(* Logix 5000 project; controller OWF Emulate 5570 rev 30.12; software revision 30.00 *) (continued)
   	OWF_Key[105,2]:=1079186439;
   	OWF_Key[105,3]:=354175718;
   	OWF_Key[105,4]:=460014900;
   	OWF_Key[105,5]:=657327792;
   	OWF_Key[105,6]:=1238184223;
   	OWF_Key[105,7]:=613398807;
   	OWF_Key[105,8]:=313681701;
   	OWF_Key[106,0]:=623677644;
   	OWF_Key[106,1]:=1206586343;
   	OWF_Key[106,2]:=1211299162;
   	OWF_Key[106,3]:=1368157030;
   	OWF_Key[106,4]:=1726692177;
   	OWF_Key[106,5]:=909079139;
   	OWF_Key[106,6]:=1189133566;
   	OWF_Key[106,7]:=1775183384;
   	OWF_Key[106,8]:=1947314078;
   	OWF_Key[107,0]:=795842741;
   	OWF_Key[107,1]:=5243211;
   	OWF_Key[107,2]:=2117485737;
   	OWF_Key[107,3]:=1222955765;
   	OWF_Key[107,4]:=1010466652;
   	OWF_Key[107,5]:=1366757084;
   	OWF_Key[107,6]:=1745897474;
   	OWF_Key[107,7]:=1196628900;
   	OWF_Key[107,8]:=422811900;
   	OWF_Key[108,0]:=51546250;
   	OWF_Key[108,1]:=1371654065;
   	OWF_Key[108,2]:=594730613;
   	OWF_Key[108,3]:=1178928938;
   	OWF_Key[108,4]:=19658574;
   	OWF_Key[108,5]:=44268080;
   	OWF_Key[108,6]:=1705061822;
   	OWF_Key[108,7]:=765733996;
   	OWF_Key[108,8]:=254021521;
   	OWF_Key[109,0]:=1089931182;
   	OWF_Key[109,1]:=456261576;
   	OWF_Key[109,2]:=1032396223;
   	OWF_Key[109,3]:=1215239566;
   	OWF_Key[109,4]:=1432021362;
   	OWF_Key[109,5]:=1482695855;
   	OWF_Key[109,6]:=471826292;
   	OWF_Key[109,7]:=1639233209;
   	OWF_Key[109,8]:=33522508;
   	OWF_Key[110,0]:=1943548851;
   	OWF_Key[110,1]:=188222712;
   	OWF_Key[110,2]:=2073166455;
   	OWF_Key[110,3]:=1482931688;
   	OWF_Key[110,4]:=816300030;
   	OWF_Key[110,5]:=246963335;
   	OWF_Key[110,6]:=313723350;
   	OWF_Key[110,7]:=331932254;
   	OWF_Key[110,8]:=1039085928;
   	OWF_Key[111,0]:=913532003;
   	OWF_Key[111,1]:=1339665160;
   	OWF_Key[111,2]:=14150618;
   	OWF_Key[111,3]:=743204030;
   	OWF_Key[111,4]:=2083710274;
   	OWF_Key[111,5]:=1872451661;
   	OWF_Key[111,6]:=1349153003;
   	OWF_Key[111,7]:=373058060;
   	OWF_Key[111,8]:=778338392;
   	OWF_Key[112,0]:=1413062923;
   	OWF_Key[112,1]:=1525503190;
   	OWF_Key[112,2]:=153669953;
   	OWF_Key[112,3]:=1075488387;
   	OWF_Key[112,4]:=1611202824;
   	OWF_Key[112,5]:=842678039;
   	OWF_Key[112,6]:=1878241110;
   	OWF_Key[112,7]:=2094622845;
   	OWF_Key[112,8]:=346061363;
   	OWF_Key[113,0]:=2007662486;
   	OWF_Key[113,1]:=609926961;
   	OWF_Key[113,2]:=208768431;
   	OWF_Key[113,3]:=1089775410;
   	OWF_Key[113,4]:=2139360128;
   	OWF_Key[113,5]:=246842036;
   	OWF_Key[113,6]:=437887573;
   	OWF_Key[113,7]:=1715106097;
   	OWF_Key[113,8]:=1931243001;
   	OWF_Key[114,0]:=1695412974;
   	OWF_Key[114,1]:=75402688;
   	OWF_Key[114,2]:=1324107774;
   	OWF_Key[114,3]:=1762126149;
   	OWF_Key[114,4]:=2045453401;
   	OWF_Key[114,5]:=1322782179;
   	OWF_Key[114,6]:=560014314;
   	OWF_Key[114,7]:=113230679;
   	OWF_Key[114,8]:=1460013455;
   	OWF_Key[115,0]:=1522550142;
   	OWF_Key[115,1]:=181079064;
   	OWF_Key[115,2]:=1318356612;
   	OWF_Key[115,3]:=1089396761;
   	OWF_Key[115,4]:=2100774490;
   	OWF_Key[115,5]:=1187593175;
   	OWF_Key[115,6]:=673723015;
   	OWF_Key[115,7]:=1625716407;
   	OWF_Key[115,8]:=157879385;
   	OWF_Key[116,0]:=1574439302;
   	OWF_Key[116,1]:=1171649064;
   	OWF_Key[116,2]:=1725295889;
   	OWF_Key[116,3]:=1508609966;
   	OWF_Key[116,4]:=893053329;
   	OWF_Key[116,5]:=2022024439;
   	OWF_Key[116,6]:=1645938530;
   	OWF_Key[116,7]:=1690657533;
   	OWF_Key[116,8]:=1383145517;
   	OWF_Key[117,0]:=255569215;
   	OWF_Key[117,1]:=1987873809;
   	OWF_Key[117,2]:=397411303;
   	OWF_Key[117,3]:=1688889668;
   	OWF_Key[117,4]:=222285489;
   	OWF_Key[117,5]:=449962612;
   	OWF_Key[117,6]:=751498151;
   	OWF_Key[117,7]:=708509537;
   	OWF_Key[117,8]:=2068975187;
   	OWF_Key[118,0]:=755822791;
   	OWF_Key[118,1]:=705169811;
   	OWF_Key[118,2]:=1142286417;
   	OWF_Key[118,3]:=157784650;
   	OWF_Key[118,4]:=506439582;
   	OWF_Key[118,5]:=1051639190;
   	OWF_Key[118,6]:=1903419853;
   	OWF_Key[118,7]:=1851507373;
   	OWF_Key[118,8]:=1030591932;
   	OWF_Key[119,0]:=2057479898;
   	OWF_Key[119,1]:=2036906294;
   	OWF_Key[119,2]:=254059922;
   	OWF_Key[119,3]:=849168680;
   	OWF_Key[119,4]:=301288022;
   	OWF_Key[119,5]:=1586180160;
   	OWF_Key[119,6]:=434263535;
   	OWF_Key[119,7]:=1375534755;
   	OWF_Key[119,8]:=967855848;
   	OWF_Key[120,0]:=1790809297;
   	OWF_Key[120,1]:=913198018;
   	OWF_Key[120,2]:=996748500;
   	OWF_Key[120,3]:=326041118;
   	OWF_Key[120,4]:=1340890547;
   	OWF_Key[120,5]:=1923120038;
   	OWF_Key[120,6]:=122657393;
   	OWF_Key[120,7]:=1589302007;
   	OWF_Key[120,8]:=1782178774;
   	OWF_Key[121,0]:=82130336;
   	OWF_Key[121,1]:=1724730757;
   	OWF_Key[121,2]:=1991211720;
   	OWF_Key[121,3]:=559635139;
   	OWF_Key[121,4]:=1292994698;
   	OWF_Key[121,5]:=884899297;
   	OWF_Key[121,6]:=54837547;
   	OWF_Key[121,7]:=1512359967;
   	OWF_Key[121,8]:=1206990758;
   	OWF_Key[122,0]:=521842158;
   	OWF_Key[122,1]:=740641184;
   	OWF_Key[122,2]:=1937985441;
   	OWF_Key[122,3]:=1079005365;
   	OWF_Key[122,4]:=1876008654;
   	OWF_Key[122,5]:=321093037;
   	OWF_Key[122,6]:=289229113;
   	OWF_Key[122,7]:=1025583141;
   	OWF_Key[122,8]:=459288858;
   	OWF_Key[123,0]:=1974309623;
   	OWF_Key[123,1]:=6712638;
   	OWF_Key[123,2]:=2007167640;
   	OWF_Key[123,3]:=27983471;
   	OWF_Key[123,4]:=1975409524;
   	OWF_Key[123,5]:=640991423;
   	OWF_Key[123,6]:=1662465747;
   	OWF_Key[123,7]:=245495606;
   	OWF_Key[123,8]:=2018234465;
   	OWF_Key[124,0]:=2095859398;
   	OWF_Key[124,1]:=1539650695;
   	OWF_Key[124,2]:=906115698;
   	OWF_Key[124,3]:=1464160346;
   	OWF_Key[124,4]:=551406825;
   	OWF_Key[124,5]:=668952051;
   	OWF_Key[124,6]:=877137102;
   	OWF_Key[124,7]:=1537695198;
   	OWF_Key[124,8]:=980602547;
   	OWF_Key[125,0]:=867529616;
   	OWF_Key[125,1]:=1849049743;
   	OWF_Key[125,2]:=991319418;
   	OWF_Key[125,3]:=1321355899;
   	OWF_Key[125,4]:=2060073135;
   	OWF_Key[125,5]:=1331119873;
   	OWF_Key[125,6]:=573685862;
   	OWF_Key[125,7]:=120334861;
   	OWF_Key[125,8]:=1086526851;
   	OWF_Key[126,0]:=1200278151;
   	OWF_Key[126,1]:=1471285710;
   	OWF_Key[126,2]:=198401618;
   	OWF_Key[126,3]:=799880776;
   	OWF_Key[126,4]:=1720054826;
   	OWF_Key[126,5]:=1991869151;
   	OWF_Key[126,6]:=524127183;
   	OWF_Key[126,7]:=241644883;
   	OWF_Key[126,8]:=464828034;
   	OWF_Key[127,0]:=703402634;
   	OWF_Key[127,1]:=1693118228;
   	OWF_Key[127,2]:=982697312;
   	OWF_Key[127,3]:=1186000843;
   	OWF_Key[127,4]:=766837985;
   	OWF_Key[127,5]:=835588933;
   	OWF_Key[127,6]:=889769892;
   	OWF_Key[127,7]:=3971994;
   	OWF_Key[127,8]:=209421061;
   	OWF_Key[128,0]:=2095700593;
   	OWF_Key[128,1]:=990463176;
   	OWF_Key[128,2]:=1203561158;
   	OWF_Key[128,3]:=1925791782;
   	OWF_Key[128,4]:=1282291352;
   	OWF_Key[128,5]:=92788621;
   	OWF_Key[128,6]:=883679225;
   	OWF_Key[128,7]:=261939133;
   	OWF_Key[128,8]:=417337857;
   	OWF_Key[129,0]:=461069728;
   	OWF_Key[129,1]:=306980987;
   	OWF_Key[129,2]:=1642188911;
   	OWF_Key[129,3]:=1558513048;
   	OWF_Key[129,4]:=235034413;
   	OWF_Key[129,5]:=49348981;
   	OWF_Key[129,6]:=119647358;
   	OWF_Key[129,7]:=1423657742;
   	OWF_Key[129,8]:=14198199;
   	OWF_Key[130,0]:=2094498674;
   	OWF_Key[130,1]:=51839195;
   	OWF_Key[130,2]:=1281989587;
   	OWF_Key[130,3]:=1580160455;
   	OWF_Key[130,4]:=1842110844;
   	OWF_Key[130,5]:=2018159406;
   	OWF_Key[130,6]:=1939031114;
   	OWF_Key[130,7]:=78193792;
   	OWF_Key[130,8]:=1487552029;
   	OWF_Key[131,0]:=1941470018;
   	OWF_Key[131,1]:=1268445567;
   	OWF_Key[131,2]:=393960364;
   	OWF_Key[131,3]:=936797167;
   	OWF_Key[131,4]:=954420768;
   	OWF_Key[131,5]:=744806357;
   	OWF_Key[131,6]:=184261489;
   	OWF_Key[131,7]:=381311501;
   	OWF_Key[131,8]:=603469973;
   	OWF_Key[132,0]:=1850055018;
   	OWF_Key[132,1]:=1224396901;
   	OWF_Key[132,2]:=296829909;
   	OWF_Key[132,3]:=249886151;
   	OWF_Key[132,4]:=1549094132;
   	OWF_Key[132,5]:=1532416817;
   	OWF_Key[132,6]:=236336348;
   	OWF_Key[132,7]:=538644360;
   	OWF_Key[132,8]:=1083710908;
   	OWF_Key[133,0]:=348017081;
   	OWF_Key[133,1]:=56755330;
   	OWF_Key[133,2]:=556981986;
   	OWF_Key[133,3]:=1776044918;
   	OWF_Key[133,4]:=828262639;
   	OWF_Key[133,5]:=409711071;
   	OWF_Key[133,6]:=1561047683;
   	OWF_Key[133,7]:=1569038695;
   	OWF_Key[133,8]:=429996743;
   	OWF_Key[134,0]:=2112779550;
   	OWF_Key[134,1]:=1981865144;
   	OWF_Key[134,2]:=381593226;
   	OWF_Key[134,3]:=1021177217;
   	OWF_Key[134,4]:=390679611;
   	OWF_Key[134,5]:=790113723;
   	OWF_Key[134,6]:=1641724200;
   	OWF_Key[134,7]:=212093161;
   	OWF_Key[134,8]:=16305740;
   	OWF_Key[135,0]:=803108154;
   	OWF_Key[135,1]:=1020906832;
   	OWF_Key[135,2]:=1152571063;
   	OWF_Key[135,3]:=149359098;
   	OWF_Key[135,4]:=1013801504;
   	OWF_Key[135,5]:=1159912230;
   	OWF_Key[135,6]:=197066836;
   	OWF_Key[135,7]:=782386646;
   	OWF_Key[135,8]:=196344100;
   	OWF_Key[136,0]:=1851665471;
   	OWF_Key[136,1]:=1218121810;
   	OWF_Key[136,2]:=1491617484;
   	OWF_Key[136,3]:=1387004363;
   	OWF_Key[136,4]:=42035451;
   	OWF_Key[136,5]:=25480957;
   	OWF_Key[136,6]:=2117762465;
   	OWF_Key[136,7]:=1606577745;
   	OWF_Key[136,8]:=939292506;
   	OWF_Key[137,0]:=557257689;
   	OWF_Key[137,1]:=1408494659;
   	OWF_Key[137,2]:=1199491796;
   	OWF_Key[137,3]:=1105486138;
   	OWF_Key[137,4]:=1507604683;
   	OWF_Key[137,5]:=392467134;
   	OWF_Key[137,6]:=310580865;
   	OWF_Key[137,7]:=565134100;
   	OWF_Key[137,8]:=1015383797;
   	OWF_Key[138,0]:=135671045;
   	OWF_Key[138,1]:=877154257;
   	OWF_Key[138,2]:=1623745783;
   	OWF_Key[138,3]:=1368835238;
   	OWF_Key[138,4]:=1988863369;
   	OWF_Key[138,5]:=575749922;
   	OWF_Key[138,6]:=2030652526;
   	OWF_Key[138,7]:=402148410;
   	OWF_Key[138,8]:=366001488;
   	OWF_Key[139,0]:=1908687818;
   	OWF_Key[139,1]:=1513823005;
   	OWF_Key[139,2]:=1615947469;
   	OWF_Key[139,3]:=1278340394;
   	OWF_Key[139,4]:=440988635;
   	OWF_Key[139,5]:=1777972517;
   	OWF_Key[139,6]:=1386151211;
   	OWF_Key[139,7]:=245033079;
   	OWF_Key[139,8]:=2110607670;
   	OWF_Key[140,0]:=423637893;
   	OWF_Key[140,1]:=777652355;
   	OWF_Key[140,2]:=905960121;
   	OWF_Key[140,3]:=976448701;
   	OWF_Key[140,4]:=173370798;
   	OWF_Key[140,5]:=1707443541;
   	OWF_Key[140,6]:=6280813;
   	OWF_Key[140,7]:=1586570709;
   	OWF_Key[140,8]:=347949075;
   	OWF_Key[141,0]:=1419227260;
   	OWF_Key[141,1]:=2137996375;
   	OWF_Key[141,2]:=550826713;
   	OWF_Key[141,3]:=270319560;
   	OWF_Key[141,4]:=1761938779;
   	OWF_Key[141,5]:=1769319179;
   	OWF_Key[141,6]:=405162215;
   	OWF_Key[141,7]:=92820702;
   	OWF_Key[141,8]:=1336055719;
   	OWF_Key[142,0]:=1852175356;
   	OWF_Key[142,1]:=613281314;
   	OWF_Key[142,2]:=1990951556;
   	OWF_Key[142,3]:=872891547;
   	OWF_Key[142,4]:=953112461;
   	OWF_Key[142,5]:=981620527;
   	OWF_Key[142,6]:=1907699741;
   	OWF_Key[142,7]:=1546914583;
   	OWF_Key[142,8]:=1313804796;
   	OWF_Key[143,0]:=310065645;
   	OWF_Key[143,1]:=541527684;
   	OWF_Key[143,2]:=1794464280;
   	OWF_Key[143,3]:=2142938457;
   	OWF_Key[143,4]:=884238194;
   	OWF_Key[143,5]:=1089289658;
   	OWF_Key[143,6]:=105264285;
   	OWF_Key[143,7]:=1423736746;
   	OWF_Key[143,8]:=1615314362;
   	OWF_Key[144,0]:=6466165;
   	OWF_Key[144,1]:=1699153526;
   	OWF_Key[144,2]:=767510287;
   	OWF_Key[144,3]:=1991118986;
   	OWF_Key[144,4]:=993722231;
   	OWF_Key[144,5]:=860308270;
   	OWF_Key[144,6]:=158856948;
   	OWF_Key[144,7]:=1427057850;
   	OWF_Key[144,8]:=4852541;
   	OWF_Key[145,0]:=114049283;
   	OWF_Key[145,1]:=340164911;
   	OWF_Key[145,2]:=1299158042;
   	OWF_Key[145,3]:=980847215;
   	OWF_Key[145,4]:=244504658;
   	OWF_Key[145,5]:=958977783;
   	OWF_Key[145,6]:=2135350412;
   	OWF_Key[145,7]:=909397507;
   	OWF_Key[145,8]:=2117256790;
   	OWF_Key[146,0]:=1934900029;
   	OWF_Key[146,1]:=156617846;
   	OWF_Key[146,2]:=1371795333;
   	OWF_Key[146,3]:=1366540458;
   	OWF_Key[146,4]:=48687158;
   	OWF_Key[146,5]:=1269845503;
   	OWF_Key[146,6]:=8307368;
   	OWF_Key[146,7]:=107307532;
   	OWF_Key[146,8]:=1897257661;
   	OWF_Key[147,0]:=1879357039;
   	OWF_Key[147,1]:=47802923;
   	OWF_Key[147,2]:=1541728788;
   	OWF_Key[147,3]:=2117668139;
   	OWF_Key[147,4]:=156416501;
   	OWF_Key[147,5]:=1715571310;
   	OWF_Key[147,6]:=1519749230;
   	OWF_Key[147,7]:=2099970770;
   	OWF_Key[147,8]:=1975760820;
   	OWF_Key[148,0]:=1852780784;
   	OWF_Key[148,1]:=38176153;
   	OWF_Key[148,2]:=423887200;
   	OWF_Key[148,3]:=1438176481;
   	OWF_Key[148,4]:=924616536;
   	OWF_Key[148,5]:=788838277;
   	OWF_Key[148,6]:=1398249766;
   	OWF_Key[148,7]:=1931406790;
   	OWF_Key[148,8]:=547521605;
   	OWF_Key[149,0]:=310483879;
   	OWF_Key[149,1]:=2044864337;
   	OWF_Key[149,2]:=2074745032;
   	OWF_Key[149,3]:=218312227;
   	OWF_Key[149,4]:=663358293;
   	OWF_Key[149,5]:=1008911891;
   	OWF_Key[149,6]:=88362942;
   	OWF_Key[149,7]:=1110396514;
   	OWF_Key[149,8]:=360154673;
   	OWF_Key[150,0]:=881826593;
   	OWF_Key[150,1]:=832451696;
   	OWF_Key[150,2]:=445991601;
   	OWF_Key[150,3]:=759796708;
   	OWF_Key[150,4]:=476997475;
   	OWF_Key[150,5]:=1183502621;
   	OWF_Key[150,6]:=916489561;
   	OWF_Key[150,7]:=510673143;
   	OWF_Key[150,8]:=1442115105;
   	OWF_Key[151,0]:=2079182206;
   	OWF_Key[151,1]:=1432083559;
   	OWF_Key[151,2]:=1691672759;
   	OWF_Key[151,3]:=344070256;
   	OWF_Key[151,4]:=1226544908;
   	OWF_Key[151,5]:=156607441;
   	OWF_Key[151,6]:=1643261836;
   	OWF_Key[151,7]:=2034004198;
   	OWF_Key[151,8]:=1567782810;
   	OWF_Key[152,0]:=1850603654;
   	OWF_Key[152,1]:=546531556;
   	OWF_Key[152,2]:=86932976;
   	OWF_Key[152,3]:=2141177608;
   	OWF_Key[152,4]:=564196549;
   	OWF_Key[152,5]:=835284922;
   	OWF_Key[152,6]:=1800632995;
   	OWF_Key[152,7]:=1774044670;
   	OWF_Key[152,8]:=599227861;
   	OWF_Key[153,0]:=1126180833;
   	OWF_Key[153,1]:=537648723;
   	OWF_Key[153,2]:=2018957043;
   	OWF_Key[153,3]:=113936735;
   	OWF_Key[153,4]:=531103137;
   	OWF_Key[153,5]:=1993941201;
   	OWF_Key[153,6]:=413134648;
   	OWF_Key[153,7]:=1164000897;
   	OWF_Key[153,8]:=1238012941;
   	OWF_Key[154,0]:=295408796;
   	OWF_Key[154,1]:=1849833269;
   	OWF_Key[154,2]:=1760932004;
   	OWF_Key[154,3]:=1994788816;
   	OWF_Key[154,4]:=334968226;
   	OWF_Key[154,5]:=1335189981;
   	OWF_Key[154,6]:=1030897726;
   	OWF_Key[154,7]:=98484120;
   	OWF_Key[154,8]:=476690948;
   	OWF_Key[155,0]:=1508241687;
   	OWF_Key[155,1]:=2079350902;
   	OWF_Key[155,2]:=86726812;
   	OWF_Key[155,3]:=1399994932;
   	OWF_Key[155,4]:=1772290692;
   	OWF_Key[155,5]:=1114819488;
   	OWF_Key[155,6]:=1835301313;
   	OWF_Key[155,7]:=1280737427;
   	OWF_Key[155,8]:=1824630929;
   	OWF_Key[156,0]:=896783386;
   	OWF_Key[156,1]:=1238520221;
   	OWF_Key[156,2]:=1303521043;
   	OWF_Key[156,3]:=2000272664;
   	OWF_Key[156,4]:=1411479205;
   	OWF_Key[156,5]:=1008892499;
   	OWF_Key[156,6]:=484998019;
   	OWF_Key[156,7]:=1953304996;
   	OWF_Key[156,8]:=682024064;
   	OWF_Key[157,0]:=771714846;
   	OWF_Key[157,1]:=81580456;
   	OWF_Key[157,2]:=1440045283;
   	OWF_Key[157,3]:=2100578838;
   	OWF_Key[157,4]:=476487452;
   	OWF_Key[157,5]:=837040200;
   	OWF_Key[157,6]:=2006065241;
   	OWF_Key[157,7]:=479466024;
   	OWF_Key[157,8]:=778174154;
   	OWF_Key[158,0]:=2059881513;
   	OWF_Key[158,1]:=1267448579;
   	OWF_Key[158,2]:=1916576462;
   	OWF_Key[158,3]:=1994723050;
   	OWF_Key[158,4]:=820419189;
   	OWF_Key[158,5]:=1622629162;
   	OWF_Key[158,6]:=576842097;
   	OWF_Key[158,7]:=1911366754;
   	OWF_Key[158,8]:=102961831;
   	OWF_Key[159,0]:=1427392151;
   	OWF_Key[159,1]:=1514105500;
   	OWF_Key[159,2]:=660047527;
   	OWF_Key[159,3]:=1565529165;
   	OWF_Key[159,4]:=1064017653;
   	OWF_Key[159,5]:=2139487925;
   	OWF_Key[159,6]:=1011083314;
   	OWF_Key[159,7]:=1330962697;
   	OWF_Key[159,8]:=2109785053;
   	OWF_Key[160,0]:=2127475596;
   	OWF_Key[160,1]:=1734616045;
   	OWF_Key[160,2]:=1738700648;
   	OWF_Key[160,3]:=1364353381;
   	OWF_Key[160,4]:=722187677;
   	OWF_Key[160,5]:=1057094241;
   	OWF_Key[160,6]:=1890275756;
   	OWF_Key[160,7]:=1092681561;
   	OWF_Key[160,8]:=208772515;
   	OWF_Key[161,0]:=1737506979;
   	OWF_Key[161,1]:=2063008297;
   	OWF_Key[161,2]:=507714092;
   	OWF_Key[161,3]:=1843967597;
   	OWF_Key[161,4]:=1391846317;
   	OWF_Key[161,5]:=1765655187;
   	OWF_Key[161,6]:=660226964;
   	OWF_Key[161,7]:=323088634;
   	OWF_Key[161,8]:=1524147629;
   	OWF_Key[162,0]:=251751109;
   	OWF_Key[162,1]:=1306151556;
   	OWF_Key[162,2]:=1640455428;
   	OWF_Key[162,3]:=911639531;
   	OWF_Key[162,4]:=416058562;
   	OWF_Key[162,5]:=1465765880;
   	OWF_Key[162,6]:=725171561;
   	OWF_Key[162,7]:=1922900838;
   	OWF_Key[162,8]:=724666186;
   	OWF_Key[163,0]:=1220369580;
   	OWF_Key[163,1]:=1947739025;
   	OWF_Key[163,2]:=78159420;
   	OWF_Key[163,3]:=543101560;
   	OWF_Key[163,4]:=1829428931;
   	OWF_Key[163,5]:=109980317;
   	OWF_Key[163,6]:=12355278;
   	OWF_Key[163,7]:=1765663600;
   	OWF_Key[163,8]:=1417306458;
   	OWF_Key[164,0]:=572738398;
   	OWF_Key[164,1]:=48159729;
   	OWF_Key[164,2]:=693163862;
   	OWF_Key[164,3]:=1898500400;
   	OWF_Key[164,4]:=1571058001;
   	OWF_Key[164,5]:=4621559;
   	OWF_Key[164,6]:=449333924;
   	OWF_Key[164,7]:=1229243509;
   	OWF_Key[164,8]:=1406919702;
   	OWF_Key[165,0]:=1041036152;
   	OWF_Key[165,1]:=1280178369;
   	OWF_Key[165,2]:=637095493;
   	OWF_Key[165,3]:=1519723875;
   	OWF_Key[165,4]:=1305406659;
   	OWF_Key[165,5]:=1719036262;
   	OWF_Key[165,6]:=935798440;
   	OWF_Key[165,7]:=127819873;
   	OWF_Key[165,8]:=2080976666;
   	OWF_Key[166,0]:=195894702;
   	OWF_Key[166,1]:=259494047;
   	OWF_Key[166,2]:=513355763;
   	OWF_Key[166,3]:=216726708;
   	OWF_Key[166,4]:=1476929573;
   	OWF_Key[166,5]:=2008506606;
   	OWF_Key[166,6]:=234471157;
   	OWF_Key[166,7]:=1668706459;
   	OWF_Key[166,8]:=404547997;
   	OWF_Key[167,0]:=483956291;
   	OWF_Key[167,1]:=1224043965;
   	OWF_Key[167,2]:=1332859147;
   	OWF_Key[167,3]:=1080776045;
   	OWF_Key[167,4]:=1052501390;
   	OWF_Key[167,5]:=1070726197;
   	OWF_Key[167,6]:=774855976;
   	OWF_Key[167,7]:=974032836;
   	OWF_Key[167,8]:=738266144;
   	OWF_Key[168,0]:=1575188023;
   	OWF_Key[168,1]:=1479810340;
   	OWF_Key[168,2]:=20101954;
   	OWF_Key[168,3]:=1354372408;
   	OWF_Key[168,4]:=2109009527;
   	OWF_Key[168,5]:=792471993;
   	OWF_Key[168,6]:=178201888;
   	OWF_Key[168,7]:=1451193004;
   	OWF_Key[168,8]:=391432259;
   	OWF_Key[169,0]:=421774451;
   	OWF_Key[169,1]:=1262675059;
   	OWF_Key[169,2]:=813719905;
   	OWF_Key[169,3]:=609456596;
   	OWF_Key[169,4]:=498754612;
   	OWF_Key[169,5]:=1188467452;
   	OWF_Key[169,6]:=1182854937;
   	OWF_Key[169,7]:=659153513;
   	OWF_Key[169,8]:=273706639;
   	OWF_Key[170,0]:=1482865476;
   	OWF_Key[170,1]:=1815595385;
   	OWF_Key[170,2]:=853235449;
   	OWF_Key[170,3]:=1255526597;
   	OWF_Key[170,4]:=1621207048;
   	OWF_Key[170,5]:=221936632;
   	OWF_Key[170,6]:=1150503334;
   	OWF_Key[170,7]:=861096856;
   	OWF_Key[170,8]:=1114127009;
   	OWF_Key[171,0]:=1592480823;
   	OWF_Key[171,1]:=1399213055;
   	OWF_Key[171,2]:=1283468591;
   	OWF_Key[171,3]:=2142943148;
   	OWF_Key[171,4]:=911093767;
   	OWF_Key[171,5]:=670577402;
   	OWF_Key[171,6]:=647672518;
   	OWF_Key[171,7]:=1978288224;
   	OWF_Key[171,8]:=1724901397;
   	OWF_Key[172,0]:=1382442647;
   	OWF_Key[172,1]:=2094122618;
   	OWF_Key[172,2]:=2063357845;
   	OWF_Key[172,3]:=1215623254;
   	OWF_Key[172,4]:=1362229760;
   	OWF_Key[172,5]:=1195702408;
   	OWF_Key[172,6]:=1932516723;
   	OWF_Key[172,7]:=1247052520;
   	OWF_Key[172,8]:=161267009;
   	OWF_Key[173,0]:=882841315;
   	OWF_Key[173,1]:=865708920;
   	OWF_Key[173,2]:=214679365;
   	OWF_Key[173,3]:=1486586684;
   	OWF_Key[173,4]:=1918804195;
   	OWF_Key[173,5]:=1009714679;
   	OWF_Key[173,6]:=1253638880;
   	OWF_Key[173,7]:=379011456;
   	OWF_Key[173,8]:=1470050814;
   	OWF_Key[174,0]:=1882221522;
   	OWF_Key[174,1]:=301503457;
   	OWF_Key[174,2]:=218575431;
   	OWF_Key[174,3]:=903000683;
   	OWF_Key[174,4]:=870234460;
   	OWF_Key[174,5]:=1808326336;
   	OWF_Key[174,6]:=1256602609;
   	OWF_Key[174,7]:=2023692039;
   	OWF_Key[174,8]:=894849577;
   	OWF_Key[175,0]:=1400988581;
   	OWF_Key[175,1]:=123062937;
   	OWF_Key[175,2]:=1739425251;
   	OWF_Key[175,3]:=1096071656;
   	OWF_Key[175,4]:=220330409;
   	OWF_Key[175,5]:=155024258;
   	OWF_Key[175,6]:=1532854343;
   	OWF_Key[175,7]:=1723784427;
   	OWF_Key[175,8]:=1695723195;
   	OWF_Key[176,0]:=663225225;
   	OWF_Key[176,1]:=1273412945;
   	OWF_Key[176,2]:=645722816;
   	OWF_Key[176,3]:=596728723;
   	OWF_Key[176,4]:=881214332;
   	OWF_Key[176,5]:=1918035236;
   	OWF_Key[176,6]:=1376817636;
   	OWF_Key[176,7]:=1553944102;
   	OWF_Key[176,8]:=1374751527;
   	OWF_Key[177,0]:=1055510972;
   	OWF_Key[177,1]:=1748003753;
   	OWF_Key[177,2]:=2133375174;
   	OWF_Key[177,3]:=1845338381;
   	OWF_Key[177,4]:=1912573970;
   	OWF_Key[177,5]:=1264078779;
   	OWF_Key[177,6]:=998137387;
   	OWF_Key[177,7]:=42399117;
   	OWF_Key[177,8]:=464555364;
   	OWF_Key[178,0]:=1334686498;
   	OWF_Key[178,1]:=1499168875;
   	OWF_Key[178,2]:=1105348302;
   	OWF_Key[178,3]:=1360557853;
   	OWF_Key[178,4]:=1408369260;
   	OWF_Key[178,5]:=832022980;
   	OWF_Key[178,6]:=1530713296;
   	OWF_Key[178,7]:=1462239575;
   	OWF_Key[178,8]:=147554149;
   	OWF_Key[179,0]:=337736197;
   	OWF_Key[179,1]:=804094734;
   	OWF_Key[179,2]:=1424134994;
   	OWF_Key[179,3]:=819569551;
   	OWF_Key[179,4]:=1642760473;
   	OWF_Key[179,5]:=1250022214;
   	OWF_Key[179,6]:=1834593966;
   	OWF_Key[179,7]:=52358876;
   	OWF_Key[179,8]:=2089055339;
   	OWF_Key[180,0]:=785374353;
   	OWF_Key[180,1]:=1851192545;
   	OWF_Key[180,2]:=546911890;
   	OWF_Key[180,3]:=294834869;
   	OWF_Key[180,4]:=149284009;
   	OWF_Key[180,5]:=1228272309;
   	OWF_Key[180,6]:=826715884;
   	OWF_Key[180,7]:=1706320570;
   	OWF_Key[180,8]:=1766167982;
   	OWF_Key[181,0]:=508304423;
   	OWF_Key[181,1]:=1081379609;
   	OWF_Key[181,2]:=1290841053;
   	OWF_Key[181,3]:=1700808611;
   	OWF_Key[181,4]:=1466979451;
   	OWF_Key[181,5]:=1772048720;
   	OWF_Key[181,6]:=294442659;
   	OWF_Key[181,7]:=476473887;
   	OWF_Key[181,8]:=312627392;
   	OWF_Key[182,0]:=130799092;
   	OWF_Key[182,1]:=370754347;
   	OWF_Key[182,2]:=490618570;
   	OWF_Key[182,3]:=1762641716;
   	OWF_Key[182,4]:=1596493207;
   	OWF_Key[182,5]:=2124642446;
   	OWF_Key[182,6]:=1488570149;
   	OWF_Key[182,7]:=487249499;
   	OWF_Key[182,8]:=2044011200;
   	OWF_Key[183,0]:=1613644728;
   	OWF_Key[183,1]:=1432050578;
   	OWF_Key[183,2]:=29955535;
   	OWF_Key[183,3]:=476437054;
   	OWF_Key[183,4]:=2071627015;
   	OWF_Key[183,5]:=1360204888;
   	OWF_Key[183,6]:=1602949651;
   	OWF_Key[183,7]:=540750401;
   	OWF_Key[183,8]:=2006341816;
   	OWF_Key[184,0]:=1863596229;
   	OWF_Key[184,1]:=1679817495;
   	OWF_Key[184,2]:=437316524;
   	OWF_Key[184,3]:=945840630;
   	OWF_Key[184,4]:=689380685;
   	OWF_Key[184,5]:=1399704068;
   	OWF_Key[184,6]:=1969338363;
   	OWF_Key[184,7]:=1138740302;
   	OWF_Key[184,8]:=1326183616;
   	OWF_Key[185,0]:=1061390855;
   	OWF_Key[185,1]:=563803020;
   	OWF_Key[185,2]:=83884656;
   	OWF_Key[185,3]:=1039791782;
   	OWF_Key[185,4]:=817193751;
   	OWF_Key[185,5]:=1967237225;
   	OWF_Key[185,6]:=206114277;
   	OWF_Key[185,7]:=2068246064;
   	OWF_Key[185,8]:=683034397;
   	OWF_Key[186,0]:=927160111;
   	OWF_Key[186,1]:=1123630525;
   	OWF_Key[186,2]:=950158315;
   	OWF_Key[186,3]:=1514936086;
   	OWF_Key[186,4]:=1183846516;
   	OWF_Key[186,5]:=849618603;
   	OWF_Key[186,6]:=920146576;
   	OWF_Key[186,7]:=2077134640;
   	OWF_Key[186,8]:=1514379988;
   	OWF_Key[187,0]:=443651777;
   	OWF_Key[187,1]:=2132346462;
   	OWF_Key[187,2]:=1651559095;
   	OWF_Key[187,3]:=2017854819;
   	OWF_Key[187,4]:=563603354;
   	OWF_Key[187,5]:=16174606;
   	OWF_Key[187,6]:=1914583408;
   	OWF_Key[187,7]:=77829821;
   	OWF_Key[187,8]:=2087537473;
   	OWF_Key[188,0]:=999926196;
   	OWF_Key[188,1]:=1281796829;
   	OWF_Key[188,2]:=399884160;
   	OWF_Key[188,3]:=1580143330;
   	OWF_Key[188,4]:=233222861;
   	OWF_Key[188,5]:=1494656376;
   	OWF_Key[188,6]:=833159469;
   	OWF_Key[188,7]:=1613980843;
   	OWF_Key[188,8]:=892065318;
   	OWF_Key[189,0]:=2086001918;
   	OWF_Key[189,1]:=1328758797;
   	OWF_Key[189,2]:=1580751688;
   	OWF_Key[189,3]:=42600786;
   	OWF_Key[189,4]:=1662052783;
   	OWF_Key[189,5]:=737217305;
   	OWF_Key[189,6]:=576824981;
   	OWF_Key[189,7]:=89486793;
   	OWF_Key[189,8]:=2014977946;
   	OWF_Key[190,0]:=1115500241;
   	OWF_Key[190,1]:=1248463029;
   	OWF_Key[190,2]:=711226434;
   	OWF_Key[190,3]:=678782870;
   	OWF_Key[190,4]:=1385507982;
   	OWF_Key[190,5]:=1794452753;
   	OWF_Key[190,6]:=1422527697;
   	OWF_Key[190,7]:=1346226311;
   	OWF_Key[190,8]:=1469236857;
   	OWF_Key[191,0]:=1784606040;
   	OWF_Key[191,1]:=810743142;
   	OWF_Key[191,2]:=1621835469;
   	OWF_Key[191,3]:=352067117;
   	OWF_Key[191,4]:=522313618;
   	OWF_Key[191,5]:=762902476;
   	OWF_Key[191,6]:=21049443;
   	OWF_Key[191,7]:=1616834552;
   	OWF_Key[191,8]:=1664708680;
   	OWF_Key[192,0]:=710739303;
   	OWF_Key[192,1]:=1353918188;
   	OWF_Key[192,2]:=918570866;
   	OWF_Key[192,3]:=148575050;
   	OWF_Key[192,4]:=1738160731;
   	OWF_Key[192,5]:=50879148;
   	OWF_Key[192,6]:=781729320;
   	OWF_Key[192,7]:=283352334;
   	OWF_Key[192,8]:=1434617957;
   	OWF_Key[193,0]:=1141588772;
   	OWF_Key[193,1]:=7773171;
   	OWF_Key[193,2]:=1622295116;
   	OWF_Key[193,3]:=1403903108;
   	OWF_Key[193,4]:=41020578;
   	OWF_Key[193,5]:=494104630;
   	OWF_Key[193,6]:=1694826823;
   	OWF_Key[193,7]:=1764796764;
   	OWF_Key[193,8]:=544023111;
   	OWF_Key[194,0]:=1990039520;
   	OWF_Key[194,1]:=176502161;
   	OWF_Key[194,2]:=382342980;
   	OWF_Key[194,3]:=371884378;
   	OWF_Key[194,4]:=1715073570;
   	OWF_Key[194,5]:=817668987;
   	OWF_Key[194,6]:=168009331;
   	OWF_Key[194,7]:=1247333616;
   	OWF_Key[194,8]:=1611506005;
   	OWF_Key[195,0]:=1125828740;
   	OWF_Key[195,1]:=1505477694;
   	OWF_Key[195,2]:=1217455241;
   	OWF_Key[195,3]:=562068804;
   	OWF_Key[195,4]:=1701570736;
   	OWF_Key[195,5]:=756978757;
   	OWF_Key[195,6]:=1345301366;
   	OWF_Key[195,7]:=1439468129;
   	OWF_Key[195,8]:=21765302;
   	OWF_Key[196,0]:=1148338672;
   	OWF_Key[196,1]:=213519708;
   	OWF_Key[196,2]:=72218494;
   	OWF_Key[196,3]:=2118826639;
   	OWF_Key[196,4]:=651041387;
   	OWF_Key[196,5]:=2056019327;
   	OWF_Key[196,6]:=1184871376;
   	OWF_Key[196,7]:=560411434;
   	OWF_Key[196,8]:=997381570;
   	OWF_Key[197,0]:=1377145466;
   	OWF_Key[197,1]:=2069573571;
   	OWF_Key[197,2]:=1677564630;
   	OWF_Key[197,3]:=841470469;
   	OWF_Key[197,4]:=1974719951;
   	OWF_Key[197,5]:=1507071811;
   	OWF_Key[197,6]:=775187470;
   	OWF_Key[197,7]:=41944172;
   	OWF_Key[197,8]:=1136356953;
   	OWF_Key[198,0]:=424494746;
   	OWF_Key[198,1]:=2091756343;
   	OWF_Key[198,2]:=1042995548;
   	OWF_Key[198,3]:=849074642;
   	OWF_Key[198,4]:=1755784134;
   	OWF_Key[198,5]:=1420218082;
   	OWF_Key[198,6]:=2035052178;
   	OWF_Key[198,7]:=1697011069;
   	OWF_Key[198,8]:=21867603;
   	OWF_Key[199,0]:=841715316;
   	OWF_Key[199,1]:=1493879133;
   	OWF_Key[199,2]:=350073662;
   	OWF_Key[199,3]:=619769092;
   	OWF_Key[199,4]:=1838864915;
   	OWF_Key[199,5]:=1429245187;
   	OWF_Key[199,6]:=716147645;
   	OWF_Key[199,7]:=1432391319;
   	OWF_Key[199,8]:=1945720998;
   	OWF_Key[200,0]:=1110374121;
   	OWF_Key[200,1]:=298532089;
   	OWF_Key[200,2]:=910156662;
   	OWF_Key[200,3]:=1380219335;
   	OWF_Key[200,4]:=1922111052;
   	OWF_Key[200,5]:=1133495485;
   	OWF_Key[200,6]:=1887604870;
   	OWF_Key[200,7]:=1809368000;
   	OWF_Key[200,8]:=394786440;
   	OWF_Key[201,0]:=318136833;
   	OWF_Key[201,1]:=2027057239;
   	OWF_Key[201,2]:=569960458;
   	OWF_Key[201,3]:=2044100499;
   	OWF_Key[201,4]:=1949964411;
   	OWF_Key[201,5]:=1078960165;
   	OWF_Key[201,6]:=1190389157;
   	OWF_Key[201,7]:=932173241;
   	OWF_Key[201,8]:=437335613;
   	OWF_Key[202,0]:=1778405543;
   	OWF_Key[202,1]:=2017189200;
   	OWF_Key[202,2]:=269590365;
   	OWF_Key[202,3]:=1087142244;
   	OWF_Key[202,4]:=311028360;
   	OWF_Key[202,5]:=707098919;
   	OWF_Key[202,6]:=586953583;
   	OWF_Key[202,7]:=2079508908;
   	OWF_Key[202,8]:=1645838479;
   	OWF_Key[203,0]:=545647947;
   	OWF_Key[203,1]:=341041339;
   	OWF_Key[203,2]:=1397694041;
   	OWF_Key[203,3]:=1886443285;
   	OWF_Key[203,4]:=699947897;
   	OWF_Key[203,5]:=340484089;
   	OWF_Key[203,6]:=551792301;
   	OWF_Key[203,7]:=811993843;
   	OWF_Key[203,8]:=1114134365;
   	OWF_Key[204,0]:=1170355825;
   	OWF_Key[204,1]:=958253245;
   	OWF_Key[204,2]:=435750162;
   	OWF_Key[204,3]:=1953679453;
   	OWF_Key[204,4]:=659548386;
   	OWF_Key[204,5]:=1759520862;
   	OWF_Key[204,6]:=170497000;
   	OWF_Key[204,7]:=1671082405;
   	OWF_Key[204,8]:=956887449;
   	OWF_Key[205,0]:=795202243;
   	OWF_Key[205,1]:=949964228;
   	OWF_Key[205,2]:=1491266862;
   	OWF_Key[205,3]:=1282569481;
   	OWF_Key[205,4]:=356150473;
   	OWF_Key[205,5]:=223471294;
   	OWF_Key[205,6]:=1426515540;
   	OWF_Key[205,7]:=172295283;
   	OWF_Key[205,8]:=1592684801;
   	OWF_Key[206,0]:=141608483;
   	OWF_Key[206,1]:=219175957;
   	OWF_Key[206,2]:=1367670659;
   	OWF_Key[206,3]:=1134541707;
   	OWF_Key[206,4]:=1982515309;
   	OWF_Key[206,5]:=520881715;
   	OWF_Key[206,6]:=1389019437;
   	OWF_Key[206,7]:=1798260508;
   	OWF_Key[206,8]:=1655812776;
   	OWF_Key[207,0]:=991428436;
   	OWF_Key[207,1]:=1134897395;
   	OWF_Key[207,2]:=253065888;
   	OWF_Key[207,3]:=1797522749;
   	OWF_Key[207,4]:=1455939091;
   	OWF_Key[207,5]:=1826217061;
   	OWF_Key[207,6]:=1693398563;
   	OWF_Key[207,7]:=1427713967;
   	OWF_Key[207,8]:=1769738933;
   	OWF_Key[208,0]:=96180913;
   	OWF_Key[208,1]:=973329616;
   	OWF_Key[208,2]:=213079395;
   	OWF_Key[208,3]:=164094998;
   	OWF_Key[208,4]:=900089502;
   	OWF_Key[208,5]:=1601256053;
   	OWF_Key[208,6]:=908582766;
   	OWF_Key[208,7]:=1288879097;
   	OWF_Key[208,8]:=1519820512;
   	OWF_Key[209,0]:=129150014;
   	OWF_Key[209,1]:=227173774;
   	OWF_Key[209,2]:=1218855506;
   	OWF_Key[209,3]:=477912913;
   	OWF_Key[209,4]:=277549162;
   	OWF_Key[209,5]:=926914002;
   	OWF_Key[209,6]:=702815136;
   	OWF_Key[209,7]:=425754552;
   	OWF_Key[209,8]:=1633235412;
   	OWF_Key[210,0]:=756957639;
   	OWF_Key[210,1]:=1747277622;
   	OWF_Key[210,2]:=1515602899;
   	OWF_Key[210,3]:=865920091;
   	OWF_Key[210,4]:=1991610208;
   	OWF_Key[210,5]:=1543655299;
   	OWF_Key[210,6]:=1135844144;
   	OWF_Key[210,7]:=1114124815;
   	OWF_Key[210,8]:=1302022684;
   	OWF_Key[211,0]:=112169027;
   	OWF_Key[211,1]:=305429435;
   	OWF_Key[211,2]:=362272662;
   	OWF_Key[211,3]:=896463526;
   	OWF_Key[211,4]:=1114812470;
   	OWF_Key[211,5]:=682696900;
   	OWF_Key[211,6]:=793916747;
   	OWF_Key[211,7]:=1622560256;
   	OWF_Key[211,8]:=1738244233;
   	OWF_Key[212,0]:=1339095545;
   	OWF_Key[212,1]:=1474097216;
   	OWF_Key[212,2]:=1845015487;
   	OWF_Key[212,3]:=741496492;
   	OWF_Key[212,4]:=1560461550;
   	OWF_Key[212,5]:=678827998;
   	OWF_Key[212,6]:=273481884;
   	OWF_Key[212,7]:=124909012;
   	OWF_Key[212,8]:=1370200106;
   	OWF_Key[213,0]:=1124601512;
   	OWF_Key[213,1]:=1165405597;
   	OWF_Key[213,2]:=914927545;
   	OWF_Key[213,3]:=1285048865;
   	OWF_Key[213,4]:=37514808;
   	OWF_Key[213,5]:=652582338;
   	OWF_Key[213,6]:=1332830376;
   	OWF_Key[213,7]:=1095513767;
   	OWF_Key[213,8]:=1915616319;
   	OWF_Key[214,0]:=763059906;
   	OWF_Key[214,1]:=2010031107;
   	OWF_Key[214,2]:=950971887;
   	OWF_Key[214,3]:=1321995046;
   	OWF_Key[214,4]:=909417107;
   	OWF_Key[214,5]:=99024424;
   	OWF_Key[214,6]:=134912494;
   	OWF_Key[214,7]:=1065568669;
   	OWF_Key[214,8]:=919737743;
   	OWF_Key[215,0]:=1919735381;
   	OWF_Key[215,1]:=515786659;
   	OWF_Key[215,2]:=1069299600;
   	OWF_Key[215,3]:=112102042;
   	OWF_Key[215,4]:=704506414;
   	OWF_Key[215,5]:=544989217;
   	OWF_Key[215,6]:=474670761;
   	OWF_Key[215,7]:=1304288593;
   	OWF_Key[215,8]:=1425535519;
   	OWF_Key[216,0]:=207099294;
   	OWF_Key[216,1]:=375022195;
   	OWF_Key[216,2]:=447822407;
   	OWF_Key[216,3]:=1369489683;
   	OWF_Key[216,4]:=1720005776;
   	OWF_Key[216,5]:=853130511;
   	OWF_Key[216,6]:=621467353;
   	OWF_Key[216,7]:=65060140;
   	OWF_Key[216,8]:=579352738;
   	OWF_Key[217,0]:=922935565;
   	OWF_Key[217,1]:=1034568947;
   	OWF_Key[217,2]:=1102036107;
   	OWF_Key[217,3]:=1223625941;
   	OWF_Key[217,4]:=392394610;
   	OWF_Key[217,5]:=308823261;
   	OWF_Key[217,6]:=1730715852;
   	OWF_Key[217,7]:=1452675602;
   	OWF_Key[217,8]:=1890168005;
   	OWF_Key[218,0]:=369917782;
   	OWF_Key[218,1]:=1855730767;
   	OWF_Key[218,2]:=1802753667;
   	OWF_Key[218,3]:=540200361;
   	OWF_Key[218,4]:=1854925038;
   	OWF_Key[218,5]:=1064842745;
   	OWF_Key[218,6]:=618917128;
   	OWF_Key[218,7]:=808975524;
   	OWF_Key[218,8]:=2091067219;
   	OWF_Key[219,0]:=1518979313;
   	OWF_Key[219,1]:=1481491188;
   	OWF_Key[219,2]:=1239679839;
   	OWF_Key[219,3]:=243248637;
   	OWF_Key[219,4]:=1671351977;
   	OWF_Key[219,5]:=1361315758;
   	OWF_Key[219,6]:=1116747920;
   	OWF_Key[219,7]:=963336063;
   	OWF_Key[219,8]:=1297413795;
   	OWF_Key[220,0]:=220574154;
   	OWF_Key[220,1]:=1851066683;
   	OWF_Key[220,2]:=1756587500;
   	OWF_Key[220,3]:=191515594;
   	OWF_Key[220,4]:=1444679663;
   	OWF_Key[220,5]:=1551868316;
   	OWF_Key[220,6]:=1148114950;
   	OWF_Key[220,7]:=297793426;
   	OWF_Key[220,8]:=1932296819;
   	OWF_Key[221,0]:=1800990008;
   	OWF_Key[221,1]:=1878116623;
   	OWF_Key[221,2]:=51389751;
   	OWF_Key[221,3]:=953438651;
   	OWF_Key[221,4]:=954775685;
   	OWF_Key[221,5]:=385010457;
   	OWF_Key[221,6]:=1874076949;
   	OWF_Key[221,7]:=1918595142;
   	OWF_Key[221,8]:=1275624116;
   	OWF_Key[222,0]:=1631559631;